   		OWF_Result[4].31:=0;
   		OWF_Result[5]:=OWF_Result[5] + 263129127+OWF_Add_c;
   		OWF_Add_c.5:=OWF_Result[5].31;
   		OWF_Result[5].31:=0;
   		OWF_Result[6]:=OWF_Result[6] + 1259933343+OWF_Add_c;
   		OWF_Add_c.6:=OWF_Result[6].31;
   		OWF_Result[6].31:=0;
   		OWF_Result[7]:=OWF_Result[7] + 1026723117+OWF_Add_c;
   		OWF_Add_c.7:=OWF_Result[7].31;
   		OWF_Result[7].31:=0;
   		OWF_Result[8]:=OWF_Result[8] + 1423999399+OWF_Add_c;
   		OWF_Add_c.8:=OWF_Result[8].31;
   		OWF_Result[8].31:=0;
   	End_If;
   	If OWF_Input[7].[6] Then
   		OWF_Result[0]:=OWF_Result[0] + 1069224909+OWF_Add_c;
   		OWF_Add_c.0:=OWF_Result[0].31;
   		OWF_Result[0].31:=0;
   		OWF_Result[1]:=OWF_Result[1] + 1534942001+OWF_Add_c;
   		OWF_Add_c.1:=OWF_Result[1].31;
   		OWF_Result[1].31:=0;
   		OWF_Result[2]:=OWF_Result[2] + 2056683021+OWF_Add_c;
   		OWF_Add_c.2:=OWF_Result[2].31;
   		OWF_Result[2].31:=0;
   		OWF_Result[3]:=OWF_Result[3] + 1056347500+OWF_Add_c;
   		OWF_Add_c.3:=OWF_Result[3].31;
   		OWF_Result[3].31:=0;
   		OWF_Result[4]:=OWF_Result[4] + 944436856+OWF_Add_c;
   		OWF_Add_c.4:=OWF_Result[4].31;
   		OWF_Result[4].31:=0;
   		OWF_Result[5]:=OWF_Result[5] + 288371840+OWF_Add_c;
   		OWF_Add_c.5:=OWF_Result[5].31;
   		OWF_Result[5].31:=0;
   		OWF_Result[6]:=OWF_Result[6] + 1541197734+OWF_Add_c;
   		OWF_Add_c.6:=OWF_Result[6].31;
   		OWF_Result[6].31:=0;
   		OWF_Result[7]:=OWF_Result[7] + 945574548+OWF_Add_c;
   		OWF_Add_c.7:=OWF_Result[7].31;
   		OWF_Result[7].31:=0;
   		OWF_Result[8]:=OWF_Result[8] + 925934982+OWF_Add_c;
   		OWF_Add_c.8:=OWF_Result[8].31;
   		OWF_Result[8].31:=0;
   	End_If;
   	If OWF_Input[7].[7] Then
   		OWF_Result[0]:=OWF_Result[0] + 2027697593+OWF_Add_c;
   		OWF_Add_c.0:=OWF_Result[0].31;
   		OWF_Result[0].31:=0;
   		OWF_Result[1]:=OWF_Result[1] + 1826137534+OWF_Add_c;
   		OWF_Add_c.1:=OWF_Result[1].31;
   		OWF_Result[1].31:=0;
   		OWF_Result[2]:=OWF_Result[2] + 1291417064+OWF_Add_c;
   		OWF_Add_c.2:=OWF_Result[2].31;
   		OWF_Result[2].31:=0;
   		OWF_Result[3]:=OWF_Result[3] + 1315183552+OWF_Add_c;
   		OWF_Add_c.3:=OWF_Result[3].31;
   		OWF_Result[3].31:=0;
   		OWF_Result[4]:=OWF_Result[4] + 492557432+OWF_Add_c;
   		OWF_Add_c.4:=OWF_Result[4].31;
   		OWF_Result[4].31:=0;
   		OWF_Result[5]:=OWF_Result[5] + 618670102+OWF_Add_c;
   		OWF_Add_c.5:=OWF_Result[5].31;
   		OWF_Result[5].31:=0;
   		OWF_Result[6]:=OWF_Result[6] + 2053349736+OWF_Add_c;
   		OWF_Add_c.6:=OWF_Result[6].31;
   		OWF_Result[6].31:=0;
   		OWF_Result[7]:=OWF_Result[7] + 286016371+OWF_Add_c;
   		OWF_Add_c.7:=OWF_Result[7].31;
   		OWF_Result[7].31:=0;
   		OWF_Result[8]:=OWF_Result[8] + 34477476+OWF_Add_c;
   		OWF_Add_c.8:=OWF_Result[8].31;
   		OWF_Result[8].31:=0;
   	End_If;
   	If OWF_Input[7].[8] Then
   		OWF_Result[0]:=OWF_Result[0] + 1609993904+OWF_Add_c;
   		OWF_Add_c.0:=OWF_Result[0].31;
   		OWF_Result[0].31:=0;
   		OWF_Result[1]:=OWF_Result[1] + 285268351+OWF_Add_c;
   		OWF_Add_c.1:=OWF_Result[1].31;
   		OWF_Result[1].31:=0;
   		OWF_Result[2]:=OWF_Result[2] + 1049093750+OWF_Add_c;
   		OWF_Add_c.2:=OWF_Result[2].31;
   		OWF_Result[2].31:=0;
   		OWF_Result[3]:=OWF_Result[3] + 12994338+OWF_Add_c;
   		OWF_Add_c.3:=OWF_Result[3].31;
   		OWF_Result[3].31:=0;
   		OWF_Result[4]:=OWF_Result[4] + 1664386814+OWF_Add_c;
   		OWF_Add_c.4:=OWF_Result[4].31;
   		OWF_Result[4].31:=0;
   		OWF_Result[5]:=OWF_Result[5] + 1612356757+OWF_Add_c;
   		OWF_Add_c.5:=OWF_Result[5].31;
   		OWF_Result[5].31:=0;
   		OWF_Result[6]:=OWF_Result[6] + 950446094+OWF_Add_c;
   		OWF_Add_c.6:=OWF_Result[6].31;
   		OWF_Result[6].31:=0;
   		OWF_Result[7]:=OWF_Result[7] + 766006761+OWF_Add_c;
   		OWF_Add_c.7:=OWF_Result[7].31;
   		OWF_Result[7].31:=0;
   		OWF_Result[8]:=OWF_Result[8] + 1355626236+OWF_Add_c;
   		OWF_Add_c.8:=OWF_Result[8].31;
   		OWF_Result[8].31:=0;
   	End_If;
   	If OWF_Input[7].[9] Then
   		OWF_Result[0]:=OWF_Result[0] + 694616675+OWF_Add_c;
   		OWF_Add_c.0:=OWF_Result[0].31;
   		OWF_Result[0].31:=0;
   		OWF_Result[1]:=OWF_Result[1] + 1636383722+OWF_Add_c;
   		OWF_Add_c.1:=OWF_Result[1].31;
   		OWF_Result[1].31:=0;
   		OWF_Result[2]:=OWF_Result[2] + 813808724+OWF_Add_c;
   		OWF_Add_c.2:=OWF_Result[2].31;
   		OWF_Result[2].31:=0;
   		OWF_Result[3]:=OWF_Result[3] + 1441798455+OWF_Add_c;
   		OWF_Add_c.3:=OWF_Result[3].31;
   		OWF_Result[3].31:=0;
   		OWF_Result[4]:=OWF_Result[4] + 205766012+OWF_Add_c;
   		OWF_Add_c.4:=OWF_Result[4].31;
   		OWF_Result[4].31:=0;
   		OWF_Result[5]:=OWF_Result[5] + 589639203+OWF_Add_c;
   		OWF_Add_c.5:=OWF_Result[5].31;
   		OWF_Result[5].31:=0;
   		OWF_Result[6]:=OWF_Result[6] + 1829006817+OWF_Add_c;
   		OWF_Add_c.6:=OWF_Result[6].31;
   		OWF_Result[6].31:=0;
   		OWF_Result[7]:=OWF_Result[7] + 1285210054+OWF_Add_c;
   		OWF_Add_c.7:=OWF_Result[7].31;
   		OWF_Result[7].31:=0;
   		OWF_Result[8]:=OWF_Result[8] + 152212693+OWF_Add_c;
   		OWF_Add_c.8:=OWF_Result[8].31;
   		OWF_Result[8].31:=0;
   	End_If;
   	If OWF_Input[7].[10] Then
   		OWF_Result[0]:=OWF_Result[0] + 306590462+OWF_Add_c;
   		OWF_Add_c.0:=OWF_Result[0].31;
   		OWF_Result[0].31:=0;
   		OWF_Result[1]:=OWF_Result[1] + 463214707+OWF_Add_c;
   		OWF_Add_c.1:=OWF_Result[1].31;
   		OWF_Result[1].31:=0;
   		OWF_Result[2]:=OWF_Result[2] + 1073243492+OWF_Add_c;
   		OWF_Add_c.2:=OWF_Result[2].31;
   		OWF_Result[2].31:=0;
   		OWF_Result[3]:=OWF_Result[3] + 1498408871+OWF_Add_c;
   		OWF_Add_c.3:=OWF_Result[3].31;
   		OWF_Result[3].31:=0;
   		OWF_Result[4]:=OWF_Result[4] + 1121005884+OWF_Add_c;
   		OWF_Add_c.4:=OWF_Result[4].31;
   		OWF_Result[4].31:=0;
   		OWF_Result[5]:=OWF_Result[5] + 1933284086+OWF_Add_c;
   		OWF_Add_c.5:=OWF_Result[5].31;
   		OWF_Result[5].31:=0;
   		OWF_Result[6]:=OWF_Result[6] + 1141991459+OWF_Add_c;
   		OWF_Add_c.6:=OWF_Result[6].31;
   		OWF_Result[6].31:=0;
   		OWF_Result[7]:=OWF_Result[7] + 1146716215+OWF_Add_c;
   		OWF_Add_c.7:=OWF_Result[7].31;
   		OWF_Result[7].31:=0;
   		OWF_Result[8]:=OWF_Result[8] + 1107820603+OWF_Add_c;
   		OWF_Add_c.8:=OWF_Result[8].31;
   		OWF_Result[8].31:=0;
   	End_If;
   	If OWF_Input[7].[11] Then
   		OWF_Result[0]:=OWF_Result[0] + 512819892+OWF_Add_c;
   		OWF_Add_c.0:=OWF_Result[0].31;
   		OWF_Result[0].31:=0;
   		OWF_Result[1]:=OWF_Result[1] + 23616385+OWF_Add_c;
   		OWF_Add_c.1:=OWF_Result[1].31;
   		OWF_Result[1].31:=0;
   		OWF_Result[2]:=OWF_Result[2] + 917671887+OWF_Add_c;
   		OWF_Add_c.2:=OWF_Result[2].31;
   		OWF_Result[2].31:=0;
   		OWF_Result[3]:=OWF_Result[3] + 355867720+OWF_Add_c;
   		OWF_Add_c.3:=OWF_Result[3].31;
   		OWF_Result[3].31:=0;
   		OWF_Result[4]:=OWF_Result[4] + 1478009650+OWF_Add_c;
   		OWF_Add_c.4:=OWF_Result[4].31;
   		OWF_Result[4].31:=0;
   		OWF_Result[5]:=OWF_Result[5] + 1568264334+OWF_Add_c;
   		OWF_Add_c.5:=OWF_Result[5].31;
   		OWF_Result[5].31:=0;
   		OWF_Result[6]:=OWF_Result[6] + 1184924613+OWF_Add_c;
   		OWF_Add_c.6:=OWF_Result[6].31;
   		OWF_Result[6].31:=0;
   		OWF_Result[7]:=OWF_Result[7] + 1527868064+OWF_Add_c;
   		OWF_Add_c.7:=OWF_Result[7].31;
   		OWF_Result[7].31:=0;
   		OWF_Result[8]:=OWF_Result[8] + 2072058158+OWF_Add_c;
   		OWF_Add_c.8:=OWF_Result[8].31;
   		OWF_Result[8].31:=0;
   	End_If;
   	If OWF_Input[7].[12] Then
   		OWF_Result[0]:=OWF_Result[0] + 1014625951+OWF_Add_c;
   		OWF_Add_c.0:=OWF_Result[0].31;
   		OWF_Result[0].31:=0;
   		OWF_Result[1]:=OWF_Result[1] + 1533249236+OWF_Add_c;
   		OWF_Add_c.1:=OWF_Result[1].31;
   		OWF_Result[1].31:=0;
   		OWF_Result[2]:=OWF_Result[2] + 2130006381+OWF_Add_c;
   		OWF_Add_c.2:=OWF_Result[2].31;
   		OWF_Result[2].31:=0;
   		OWF_Result[3]:=OWF_Result[3] + 2146846276+OWF_Add_c;
   		OWF_Add_c.3:=OWF_Result[3].31;
   		OWF_Result[3].31:=0;
   		OWF_Result[4]:=OWF_Result[4] + 1646388285+OWF_Add_c;
   		OWF_Add_c.4:=OWF_Result[4].31;
   		OWF_Result[4].31:=0;
   		OWF_Result[5]:=OWF_Result[5] + 1699246205+OWF_Add_c;
   		OWF_Add_c.5:=OWF_Result[5].31;
   		OWF_Result[5].31:=0;
   		OWF_Result[6]:=OWF_Result[6] + 559380684+OWF_Add_c;
   		OWF_Add_c.6:=OWF_Result[6].31;
   		OWF_Result[6].31:=0;
   		OWF_Result[7]:=OWF_Result[7] + 1307307102+OWF_Add_c;
   		OWF_Add_c.7:=OWF_Result[7].31;
   		OWF_Result[7].31:=0;
   		OWF_Result[8]:=OWF_Result[8] + 606704531+OWF_Add_c;
   		OWF_Add_c.8:=OWF_Result[8].31;
   		OWF_Result[8].31:=0;
   	End_If;
   	If OWF_Input[7].[13] Then
   		OWF_Result[0]:=OWF_Result[0] + 1359161121+OWF_Add_c;
   		OWF_Add_c.0:=OWF_Result[0].31;
   		OWF_Result[0].31:=0;
   		OWF_Result[1]:=OWF_Result[1] + 1918952380+OWF_Add_c;
   		OWF_Add_c.1:=OWF_Result[1].31;
   		OWF_Result[1].31:=0;
   		OWF_Result[2]:=OWF_Result[2] + 1473068338+OWF_Add_c;
   		OWF_Add_c.2:=OWF_Result[2].31;
   		OWF_Result[2].31:=0;
   		OWF_Result[3]:=OWF_Result[3] + 1693090892+OWF_Add_c;
   		OWF_Add_c.3:=OWF_Result[3].31;
   		OWF_Result[3].31:=0;
   		OWF_Result[4]:=OWF_Result[4] + 1915525502+OWF_Add_c;
   		OWF_Add_c.4:=OWF_Result[4].31;
   		OWF_Result[4].31:=0;
   		OWF_Result[5]:=OWF_Result[5] + 1372317013+OWF_Add_c;
   		OWF_Add_c.5:=OWF_Result[5].31;
   		OWF_Result[5].31:=0;
   		OWF_Result[6]:=OWF_Result[6] + 99771102+OWF_Add_c;
   		OWF_Add_c.6:=OWF_Result[6].31;
   		OWF_Result[6].31:=0;
   		OWF_Result[7]:=OWF_Result[7] + 192894431+OWF_Add_c;
   		OWF_Add_c.7:=OWF_Result[7].31;
   		OWF_Result[7].31:=0;
   		OWF_Result[8]:=OWF_Result[8] + 1744731961+OWF_Add_c;
   		OWF_Add_c.8:=OWF_Result[8].31;
   		OWF_Result[8].31:=0;
   	End_If;
   	If OWF_Input[7].[14] Then
   		OWF_Result[0]:=OWF_Result[0] + 1706736508+OWF_Add_c;
   		OWF_Add_c.0:=OWF_Result[0].31;
   		OWF_Result[0].31:=0;
   		OWF_Result[1]:=OWF_Result[1] + 1484877150+OWF_Add_c;
   		OWF_Add_c.1:=OWF_Result[1].31;
   		OWF_Result[1].31:=0;
   		OWF_Result[2]:=OWF_Result[2] + 869604235+OWF_Add_c;
   		OWF_Add_c.2:=OWF_Result[2].31;
   		OWF_Result[2].31:=0;
   		OWF_Result[3]:=OWF_Result[3] + 1353356392+OWF_Add_c;
   		OWF_Add_c.3:=OWF_Result[3].31;
   		OWF_Result[3].31:=0;
   		OWF_Result[4]:=OWF_Result[4] + 347447568+OWF_Add_c;
   		OWF_Add_c.4:=OWF_Result[4].31;
   		OWF_Result[4].31:=0;
   		OWF_Result[5]:=OWF_Result[5] + 1293208581+OWF_Add_c;
   		OWF_Add_c.5:=OWF_Result[5].31;
   		OWF_Result[5].31:=0;
   		OWF_Result[6]:=OWF_Result[6] + 1575776397+OWF_Add_c;
   		OWF_Add_c.6:=OWF_Result[6].31;
   		OWF_Result[6].31:=0;
   		OWF_Result[7]:=OWF_Result[7] + 1427687325+OWF_Add_c;
   		OWF_Add_c.7:=OWF_Result[7].31;
   		OWF_Result[7].31:=0;
   		OWF_Result[8]:=OWF_Result[8] + 935165463+OWF_Add_c;
   		OWF_Add_c.8:=OWF_Result[8].31;
   		OWF_Result[8].31:=0;
   	End_If;
   	If OWF_Input[7].[15] Then
   		OWF_Result[0]:=OWF_Result[0] + 1743664197+OWF_Add_c;
   		OWF_Add_c.0:=OWF_Result[0].31;
   		OWF_Result[0].31:=0;
   		OWF_Result[1]:=OWF_Result[1] + 706528617+OWF_Add_c;
   		OWF_Add_c.1:=OWF_Result[1].31;
   		OWF_Result[1].31:=0;
   		OWF_Result[2]:=OWF_Result[2] + 1958351723+OWF_Add_c;
   		OWF_Add_c.2:=OWF_Result[2].31;
   		OWF_Result[2].31:=0;
   		OWF_Result[3]:=OWF_Result[3] + 82257141+OWF_Add_c;
   		OWF_Add_c.3:=OWF_Result[3].31;
   		OWF_Result[3].31:=0;
   		OWF_Result[4]:=OWF_Result[4] + 860284908+OWF_Add_c;
   		OWF_Add_c.4:=OWF_Result[4].31;
   		OWF_Result[4].31:=0;
   		OWF_Result[5]:=OWF_Result[5] + 1587356663+OWF_Add_c;
   		OWF_Add_c.5:=OWF_Result[5].31;
   		OWF_Result[5].31:=0;
   		OWF_Result[6]:=OWF_Result[6] + 1299103155+OWF_Add_c;
   		OWF_Add_c.6:=OWF_Result[6].31;
   		OWF_Result[6].31:=0;
   		OWF_Result[7]:=OWF_Result[7] + 1945550030+OWF_Add_c;
   		OWF_Add_c.7:=OWF_Result[7].31;
   		OWF_Result[7].31:=0;
   		OWF_Result[8]:=OWF_Result[8] + 2117411835+OWF_Add_c;
   		OWF_Add_c.8:=OWF_Result[8].31;
   		OWF_Result[8].31:=0;
   	End_If;
   	If OWF_Input[7].[16] Then
   		OWF_Result[0]:=OWF_Result[0] + 1713469729+OWF_Add_c;
   		OWF_Add_c.0:=OWF_Result[0].31;
   		OWF_Result[0].31:=0;
   		OWF_Result[1]:=OWF_Result[1] + 581994065+OWF_Add_c;
   		OWF_Add_c.1:=OWF_Result[1].31;
   		OWF_Result[1].31:=0;
   		OWF_Result[2]:=OWF_Result[2] + 190604491+OWF_Add_c;
   		OWF_Add_c.2:=OWF_Result[2].31;
   		OWF_Result[2].31:=0;
   		OWF_Result[3]:=OWF_Result[3] + 1975804182+OWF_Add_c;
   		OWF_Add_c.3:=OWF_Result[3].31;
   		OWF_Result[3].31:=0;
   		OWF_Result[4]:=OWF_Result[4] + 1579426154+OWF_Add_c;
   		OWF_Add_c.4:=OWF_Result[4].31;
   		OWF_Result[4].31:=0;
   		OWF_Result[5]:=OWF_Result[5] + 1526883195+OWF_Add_c;
   		OWF_Add_c.5:=OWF_Result[5].31;
   		OWF_Result[5].31:=0;
   		OWF_Result[6]:=OWF_Result[6] + 1534112395+OWF_Add_c;
   		OWF_Add_c.6:=OWF_Result[6].31;
   		OWF_Result[6].31:=0;
   		OWF_Result[7]:=OWF_Result[7] + 1953195996+OWF_Add_c;
   		OWF_Add_c.7:=OWF_Result[7].31;
   		OWF_Result[7].31:=0;
   		OWF_Result[8]:=OWF_Result[8] + 1196776541+OWF_Add_c;
   		OWF_Add_c.8:=OWF_Result[8].31;
   		OWF_Result[8].31:=0;
   	End_If;
   	If OWF_Input[7].[17] Then
   		OWF_Result[0]:=OWF_Result[0] + 1352341478+OWF_Add_c;
   		OWF_Add_c.0:=OWF_Result[0].31;
   		OWF_Result[0].31:=0;
   		OWF_Result[1]:=OWF_Result[1] + 1327190218+OWF_Add_c;
   		OWF_Add_c.1:=OWF_Result[1].31;
   		OWF_Result[1].31:=0;
   		OWF_Result[2]:=OWF_Result[2] + 1940036231+OWF_Add_c;
   		OWF_Add_c.2:=OWF_Result[2].31;
   		OWF_Result[2].31:=0;
   		OWF_Result[3]:=OWF_Result[3] + 569828080+OWF_Add_c;
   		OWF_Add_c.3:=OWF_Result[3].31;
   		OWF_Result[3].31:=0;
   		OWF_Result[4]:=OWF_Result[4] + 1243727683+OWF_Add_c;
   		OWF_Add_c.4:=OWF_Result[4].31;
   		OWF_Result[4].31:=0;
   		OWF_Result[5]:=OWF_Result[5] + 741960146+OWF_Add_c;
   		OWF_Add_c.5:=OWF_Result[5].31;
   		OWF_Result[5].31:=0;
   		OWF_Result[6]:=OWF_Result[6] + 2046665451+OWF_Add_c;
   		OWF_Add_c.6:=OWF_Result[6].31;
   		OWF_Result[6].31:=0;
   		OWF_Result[7]:=OWF_Result[7] + 482388128+OWF_Add_c;
   		OWF_Add_c.7:=OWF_Result[7].31;
   		OWF_Result[7].31:=0;
   		OWF_Result[8]:=OWF_Result[8] + 1415487699+OWF_Add_c;
   		OWF_Add_c.8:=OWF_Result[8].31;
   		OWF_Result[8].31:=0;
   	End_If;
   	If OWF_Input[7].[18] Then
   		OWF_Result[0]:=OWF_Result[0] + 419967488+OWF_Add_c;
   		OWF_Add_c.0:=OWF_Result[0].31;
   		OWF_Result[0].31:=0;
   		OWF_Result[1]:=OWF_Result[1] + 319301420+OWF_Add_c;
   		OWF_Add_c.1:=OWF_Result[1].31;
   		OWF_Result[1].31:=0;
   		OWF_Result[2]:=OWF_Result[2] + 1439251767+OWF_Add_c;
   		OWF_Add_c.2:=OWF_Result[2].31;
   		OWF_Result[2].31:=0;
   		OWF_Result[3]:=OWF_Result[3] + 159030407+OWF_Add_c;
   		OWF_Add_c.3:=OWF_Result[3].31;
   		OWF_Result[3].31:=0;
   		OWF_Result[4]:=OWF_Result[4] + 1688057992+OWF_Add_c;
   		OWF_Add_c.4:=OWF_Result[4].31;
   		OWF_Result[4].31:=0;
   		OWF_Result[5]:=OWF_Result[5] + 677856544+OWF_Add_c;
   		OWF_Add_c.5:=OWF_Result[5].31;
   		OWF_Result[5].31:=0;
   		OWF_Result[6]:=OWF_Result[6] + 1921290271+OWF_Add_c;
   		OWF_Add_c.6:=OWF_Result[6].31;
   		OWF_Result[6].31:=0;
   		OWF_Result[7]:=OWF_Result[7] + 1347176510+OWF_Add_c;
   		OWF_Add_c.7:=OWF_Result[7].31;
   		OWF_Result[7].31:=0;
   		OWF_Result[8]:=OWF_Result[8] + 1129087746+OWF_Add_c;
   		OWF_Add_c.8:=OWF_Result[8].31;
   		OWF_Result[8].31:=0;
   	End_If;
   	If OWF_Input[7].[19] Then
   		OWF_Result[0]:=OWF_Result[0] + 909989480+OWF_Add_c;
   		OWF_Add_c.0:=OWF_Result[0].31;
   		OWF_Result[0].31:=0;
   		OWF_Result[1]:=OWF_Result[1] + 70607674+OWF_Add_c;
   		OWF_Add_c.1:=OWF_Result[1].31;
   		OWF_Result[1].31:=0;
   		OWF_Result[2]:=OWF_Result[2] + 102357735+OWF_Add_c;
   		OWF_Add_c.2:=OWF_Result[2].31;
   		OWF_Result[2].31:=0;
   		OWF_Result[3]:=OWF_Result[3] + 1548947751+OWF_Add_c;
   		OWF_Add_c.3:=OWF_Result[3].31;
   		OWF_Result[3].31:=0;
   		OWF_Result[4]:=OWF_Result[4] + 1541273950+OWF_Add_c;
   		OWF_Add_c.4:=OWF_Result[4].31;
   		OWF_Result[4].31:=0;
   		OWF_Result[5]:=OWF_Result[5] + 1965581916+OWF_Add_c;
   		OWF_Add_c.5:=OWF_Result[5].31;
   		OWF_Result[5].31:=0;
   		OWF_Result[6]:=OWF_Result[6] + 714783171+OWF_Add_c;
   		OWF_Add_c.6:=OWF_Result[6].31;
   		OWF_Result[6].31:=0;
   		OWF_Result[7]:=OWF_Result[7] + 952638591+OWF_Add_c;
   		OWF_Add_c.7:=OWF_Result[7].31;
   		OWF_Result[7].31:=0;
   		OWF_Result[8]:=OWF_Result[8] + 1892750752+OWF_Add_c;
   		OWF_Add_c.8:=OWF_Result[8].31;
   		OWF_Result[8].31:=0;
   	End_If;
   	If OWF_Input[7].[20] Then
   		OWF_Result[0]:=OWF_Result[0] + 1923601846+OWF_Add_c;
   		OWF_Add_c.0:=OWF_Result[0].31;
   		OWF_Result[0].31:=0;
   		OWF_Result[1]:=OWF_Result[1] + 431367542+OWF_Add_c;
   		OWF_Add_c.1:=OWF_Result[1].31;
   		OWF_Result[1].31:=0;
   		OWF_Result[2]:=OWF_Result[2] + 812772690+OWF_Add_c;
   		OWF_Add_c.2:=OWF_Result[2].31;
   		OWF_Result[2].31:=0;
   		OWF_Result[3]:=OWF_Result[3] + 1612004830+OWF_Add_c;
   		OWF_Add_c.3:=OWF_Result[3].31;
   		OWF_Result[3].31:=0;
   		OWF_Result[4]:=OWF_Result[4] + 1503607425+OWF_Add_c;
   		OWF_Add_c.4:=OWF_Result[4].31;
   		OWF_Result[4].31:=0;
   		OWF_Result[5]:=OWF_Result[5] + 257117095+OWF_Add_c;
   		OWF_Add_c.5:=OWF_Result[5].31;
   		OWF_Result[5].31:=0;
   		OWF_Result[6]:=OWF_Result[6] + 1165565758+OWF_Add_c;
   		OWF_Add_c.6:=OWF_Result[6].31;
   		OWF_Result[6].31:=0;
   		OWF_Result[7]:=OWF_Result[7] + 1791078952+OWF_Add_c;
   		OWF_Add_c.7:=OWF_Result[7].31;
   		OWF_Result[7].31:=0;
   		OWF_Result[8]:=OWF_Result[8] + 1316586480+OWF_Add_c;
   		OWF_Add_c.8:=OWF_Result[8].31;
   		OWF_Result[8].31:=0;
   	End_If;
   	If OWF_Input[7].[21] Then
   		OWF_Result[0]:=OWF_Result[0] + 1179130031+OWF_Add_c;
   		OWF_Add_c.0:=OWF_Result[0].31;
   		OWF_Result[0].31:=0;
   		OWF_Result[1]:=OWF_Result[1] + 1413483742+OWF_Add_c;
   		OWF_Add_c.1:=OWF_Result[1].31;
   		OWF_Result[1].31:=0;
   		OWF_Result[2]:=OWF_Result[2] + 2076538493+OWF_Add_c;
   		OWF_Add_c.2:=OWF_Result[2].31;
   		OWF_Result[2].31:=0;
   		OWF_Result[3]:=OWF_Result[3] + 415974763+OWF_Add_c;
   		OWF_Add_c.3:=OWF_Result[3].31;
   		OWF_Result[3].31:=0;
   		OWF_Result[4]:=OWF_Result[4] + 461079233+OWF_Add_c;
   		OWF_Add_c.4:=OWF_Result[4].31;
   		OWF_Result[4].31:=0;
   		OWF_Result[5]:=OWF_Result[5] + 207770264+OWF_Add_c;
   		OWF_Add_c.5:=OWF_Result[5].31;
   		OWF_Result[5].31:=0;
   		OWF_Result[6]:=OWF_Result[6] + 670532004+OWF_Add_c;
   		OWF_Add_c.6:=OWF_Result[6].31;
   		OWF_Result[6].31:=0;
   		OWF_Result[7]:=OWF_Result[7] + 164283060+OWF_Add_c;
   		OWF_Add_c.7:=OWF_Result[7].31;
   		OWF_Result[7].31:=0;
   		OWF_Result[8]:=OWF_Result[8] + 1512816438+OWF_Add_c;
   		OWF_Add_c.8:=OWF_Result[8].31;
   		OWF_Result[8].31:=0;
   	End_If;
   	If OWF_Input[7].[22] Then
   		OWF_Result[0]:=OWF_Result[0] + 1897360171+OWF_Add_c;
   		OWF_Add_c.0:=OWF_Result[0].31;
   		OWF_Result[0].31:=0;
   		OWF_Result[1]:=OWF_Result[1] + 1308779824+OWF_Add_c;
   		OWF_Add_c.1:=OWF_Result[1].31;
   		OWF_Result[1].31:=0;
   		OWF_Result[2]:=OWF_Result[2] + 1875593423+OWF_Add_c;
   		OWF_Add_c.2:=OWF_Result[2].31;
   		OWF_Result[2].31:=0;
   		OWF_Result[3]:=OWF_Result[3] + 571271217+OWF_Add_c;
   		OWF_Add_c.3:=OWF_Result[3].31;
   		OWF_Result[3].31:=0;
   		OWF_Result[4]:=OWF_Result[4] + 344940971+OWF_Add_c;
   		OWF_Add_c.4:=OWF_Result[4].31;
   		OWF_Result[4].31:=0;
   		OWF_Result[5]:=OWF_Result[5] + 75339231+OWF_Add_c;
   		OWF_Add_c.5:=OWF_Result[5].31;
   		OWF_Result[5].31:=0;
   		OWF_Result[6]:=OWF_Result[6] + 1428316860+OWF_Add_c;
   		OWF_Add_c.6:=OWF_Result[6].31;
   		OWF_Result[6].31:=0;
   		OWF_Result[7]:=OWF_Result[7] + 1811603075+OWF_Add_c;
   		OWF_Add_c.7:=OWF_Result[7].31;
   		OWF_Result[7].31:=0;
   		OWF_Result[8]:=OWF_Result[8] + 1679786029+OWF_Add_c;
   		OWF_Add_c.8:=OWF_Result[8].31;
   		OWF_Result[8].31:=0;
   	End_If;
   	If OWF_Input[7].[23] Then
   		OWF_Result[0]:=OWF_Result[0] + 271831917+OWF_Add_c;
   		OWF_Add_c.0:=OWF_Result[0].31;
   		OWF_Result[0].31:=0;
   		OWF_Result[1]:=OWF_Result[1] + 663117307+OWF_Add_c;
   		OWF_Add_c.1:=OWF_Result[1].31;
   		OWF_Result[1].31:=0;
   		OWF_Result[2]:=OWF_Result[2] + 1802435718+OWF_Add_c;
   		OWF_Add_c.2:=OWF_Result[2].31;
   		OWF_Result[2].31:=0;
   		OWF_Result[3]:=OWF_Result[3] + 585874673+OWF_Add_c;
   		OWF_Add_c.3:=OWF_Result[3].31;
   		OWF_Result[3].31:=0;
   		OWF_Result[4]:=OWF_Result[4] + 701698092+OWF_Add_c;
   		OWF_Add_c.4:=OWF_Result[4].31;
   		OWF_Result[4].31:=0;
   		OWF_Result[5]:=OWF_Result[5] + 1402770880+OWF_Add_c;
   		OWF_Add_c.5:=OWF_Result[5].31;
   		OWF_Result[5].31:=0;
   		OWF_Result[6]:=OWF_Result[6] + 452824658+OWF_Add_c;
   		OWF_Add_c.6:=OWF_Result[6].31;
   		OWF_Result[6].31:=0;
   		OWF_Result[7]:=OWF_Result[7] + 1400742763+OWF_Add_c;
   		OWF_Add_c.7:=OWF_Result[7].31;
   		OWF_Result[7].31:=0;
   		OWF_Result[8]:=OWF_Result[8] + 2073024045+OWF_Add_c;
   		OWF_Add_c.8:=OWF_Result[8].31;
   		OWF_Result[8].31:=0;
   	End_If;
   	If OWF_Input[7].[24] Then
   		OWF_Result[0]:=OWF_Result[0] + 1367845667+OWF_Add_c;
   		OWF_Add_c.0:=OWF_Result[0].31;
   		OWF_Result[0].31:=0;
   		OWF_Result[1]:=OWF_Result[1] + 1195094582+OWF_Add_c;
   		OWF_Add_c.1:=OWF_Result[1].31;
   		OWF_Result[1].31:=0;
   		OWF_Result[2]:=OWF_Result[2] + 494736933+OWF_Add_c;
   		OWF_Add_c.2:=OWF_Result[2].31;
   		OWF_Result[2].31:=0;
   		OWF_Result[3]:=OWF_Result[3] + 1875737261+OWF_Add_c;
   		OWF_Add_c.3:=OWF_Result[3].31;
   		OWF_Result[3].31:=0;
   		OWF_Result[4]:=OWF_Result[4] + 726339725+OWF_Add_c;
   		OWF_Add_c.4:=OWF_Result[4].31;
   		OWF_Result[4].31:=0;
   		OWF_Result[5]:=OWF_Result[5] + 1862851936+OWF_Add_c;
   		OWF_Add_c.5:=OWF_Result[5].31;
   		OWF_Result[5].31:=0;
   		OWF_Result[6]:=OWF_Result[6] + 296798862+OWF_Add_c;
   		OWF_Add_c.6:=OWF_Result[6].31;
   		OWF_Result[6].31:=0;
   		OWF_Result[7]:=OWF_Result[7] + 1485306441+OWF_Add_c;
   		OWF_Add_c.7:=OWF_Result[7].31;
   		OWF_Result[7].31:=0;
   		OWF_Result[8]:=OWF_Result[8] + 79244469+OWF_Add_c;
   		OWF_Add_c.8:=OWF_Result[8].31;
   		OWF_Result[8].31:=0;
   	End_If;
   	If OWF_Input[7].[25] Then
   		OWF_Result[0]:=OWF_Result[0] + 1748009068+OWF_Add_c;
   		OWF_Add_c.0:=OWF_Result[0].31;
   		OWF_Result[0].31:=0;
   		OWF_Result[1]:=OWF_Result[1] + 153673379+OWF_Add_c;
   		OWF_Add_c.1:=OWF_Result[1].31;
   		OWF_Result[1].31:=0;
   		OWF_Result[2]:=OWF_Result[2] + 1563899973+OWF_Add_c;
   		OWF_Add_c.2:=OWF_Result[2].31;
   		OWF_Result[2].31:=0;
   		OWF_Result[3]:=OWF_Result[3] + 210477071+OWF_Add_c;
   		OWF_Add_c.3:=OWF_Result[3].31;
   		OWF_Result[3].31:=0;
   		OWF_Result[4]:=OWF_Result[4] + 598591903+OWF_Add_c;
   		OWF_Add_c.4:=OWF_Result[4].31;
   		OWF_Result[4].31:=0;
   		OWF_Result[5]:=OWF_Result[5] + 889903791+OWF_Add_c;
   		OWF_Add_c.5:=OWF_Result[5].31;
   		OWF_Result[5].31:=0;
   		OWF_Result[6]:=OWF_Result[6] + 1087681228+OWF_Add_c;
   		OWF_Add_c.6:=OWF_Result[6].31;
   		OWF_Result[6].31:=0;
   		OWF_Result[7]:=OWF_Result[7] + 146945819+OWF_Add_c;
   		OWF_Add_c.7:=OWF_Result[7].31;
   		OWF_Result[7].31:=0;
   		OWF_Result[8]:=OWF_Result[8] + 658778953+OWF_Add_c;
   		OWF_Add_c.8:=OWF_Result[8].31;
   		OWF_Result[8].31:=0;
   	End_If;
   	If OWF_Input[7].[26] Then
   		OWF_Result[0]:=OWF_Result[0] + 1388889236+OWF_Add_c;
   		OWF_Add_c.0:=OWF_Result[0].31;
   		OWF_Result[0].31:=0;
   		OWF_Result[1]:=OWF_Result[1] + 1854230592+OWF_Add_c;
   		OWF_Add_c.1:=OWF_Result[1].31;
   		OWF_Result[1].31:=0;
   		OWF_Result[2]:=OWF_Result[2] + 1952659775+OWF_Add_c;
   		OWF_Add_c.2:=OWF_Result[2].31;
   		OWF_Result[2].31:=0;
   		OWF_Result[3]:=OWF_Result[3] + 693016622+OWF_Add_c;
   		OWF_Add_c.3:=OWF_Result[3].31;
   		OWF_Result[3].31:=0;
   		OWF_Result[4]:=OWF_Result[4] + 19961190+OWF_Add_c;
   		OWF_Add_c.4:=OWF_Result[4].31;
   		OWF_Result[4].31:=0;
   		OWF_Result[5]:=OWF_Result[5] + 1155238848+OWF_Add_c;
   		OWF_Add_c.5:=OWF_Result[5].31;
   		OWF_Result[5].31:=0;
   		OWF_Result[6]:=OWF_Result[6] + 1721973623+OWF_Add_c;
   		OWF_Add_c.6:=OWF_Result[6].31;
   		OWF_Result[6].31:=0;
   		OWF_Result[7]:=OWF_Result[7] + 1298626904+OWF_Add_c;
   		OWF_Add_c.7:=OWF_Result[7].31;
   		OWF_Result[7].31:=0;
   		OWF_Result[8]:=OWF_Result[8] + 704184103+OWF_Add_c;
   		OWF_Add_c.8:=OWF_Result[8].31;
   		OWF_Result[8].31:=0;
   	End_If;
   	If OWF_Input[7].[27] Then
   		OWF_Result[0]:=OWF_Result[0] + 1064559134+OWF_Add_c;
   		OWF_Add_c.0:=OWF_Result[0].31;
   		OWF_Result[0].31:=0;
   		OWF_Result[1]:=OWF_Result[1] + 628496468+OWF_Add_c;
   		OWF_Add_c.1:=OWF_Result[1].31;
   		OWF_Result[1].31:=0;
   		OWF_Result[2]:=OWF_Result[2] + 1741787667+OWF_Add_c;
   		OWF_Add_c.2:=OWF_Result[2].31;
   		OWF_Result[2].31:=0;
   		OWF_Result[3]:=OWF_Result[3] + 650880797+OWF_Add_c;
   		OWF_Add_c.3:=OWF_Result[3].31;
   		OWF_Result[3].31:=0;
   		OWF_Result[4]:=OWF_Result[4] + 927193641+OWF_Add_c;
   		OWF_Add_c.4:=OWF_Result[4].31;
   		OWF_Result[4].31:=0;
   		OWF_Result[5]:=OWF_Result[5] + 690779087+OWF_Add_c;
   		OWF_Add_c.5:=OWF_Result[5].31;
   		OWF_Result[5].31:=0;
   		OWF_Result[6]:=OWF_Result[6] + 1387171811+OWF_Add_c;
   		OWF_Add_c.6:=OWF_Result[6].31;
   		OWF_Result[6].31:=0;
   		OWF_Result[7]:=OWF_Result[7] + 1642242275+OWF_Add_c;
   		OWF_Add_c.7:=OWF_Result[7].31;
   		OWF_Result[7].31:=0;
   		OWF_Result[8]:=OWF_Result[8] + 750154437+OWF_Add_c;
   		OWF_Add_c.8:=OWF_Result[8].31;
   		OWF_Result[8].31:=0;
   	End_If;
   	If OWF_Input[7].[28] Then
   		OWF_Result[0]:=OWF_Result[0] + 1648370074+OWF_Add_c;
   		OWF_Add_c.0:=OWF_Result[0].31;
   		OWF_Result[0].31:=0;
   		OWF_Result[1]:=OWF_Result[1] + 242619355+OWF_Add_c;
   		OWF_Add_c.1:=OWF_Result[1].31;
   		OWF_Result[1].31:=0;
   		OWF_Result[2]:=OWF_Result[2] + 1874736599+OWF_Add_c;
   		OWF_Add_c.2:=OWF_Result[2].31;
   		OWF_Result[2].31:=0;
   		OWF_Result[3]:=OWF_Result[3] + 1413909693+OWF_Add_c;
   		OWF_Add_c.3:=OWF_Result[3].31;
   		OWF_Result[3].31:=0;
   		OWF_Result[4]:=OWF_Result[4] + 415302371+OWF_Add_c;
   		OWF_Add_c.4:=OWF_Result[4].31;
   		OWF_Result[4].31:=0;
   		OWF_Result[5]:=OWF_Result[5] + 2103173316+OWF_Add_c;
   		OWF_Add_c.5:=OWF_Result[5].31;
   		OWF_Result[5].31:=0;
   		OWF_Result[6]:=OWF_Result[6] + 317087375+OWF_Add_c;
   		OWF_Add_c.6:=OWF_Result[6].31;
   		OWF_Result[6].31:=0;
   		OWF_Result[7]:=OWF_Result[7] + 1550821217+OWF_Add_c;
   		OWF_Add_c.7:=OWF_Result[7].31;
   		OWF_Result[7].31:=0;
   		OWF_Result[8]:=OWF_Result[8] + 61155956+OWF_Add_c;
   		OWF_Add_c.8:=OWF_Result[8].31;
   		OWF_Result[8].31:=0;
   	End_If;
   	If OWF_Input[7].[29] Then
   		OWF_Result[0]:=OWF_Result[0] + 632604897+OWF_Add_c;
   		OWF_Add_c.0:=OWF_Result[0].31;
   		OWF_Result[0].31:=0;
   		OWF_Result[1]:=OWF_Result[1] + 1890179507+OWF_Add_c;
   		OWF_Add_c.1:=OWF_Result[1].31;
   		OWF_Result[1].31:=0;
   		OWF_Result[2]:=OWF_Result[2] + 1607995656+OWF_Add_c;
   		OWF_Add_c.2:=OWF_Result[2].31;
   		OWF_Result[2].31:=0;
   		OWF_Result[3]:=OWF_Result[3] + 1449206150+OWF_Add_c;
   		OWF_Add_c.3:=OWF_Result[3].31;
   		OWF_Result[3].31:=0;
   		OWF_Result[4]:=OWF_Result[4] + 402726737+OWF_Add_c;
   		OWF_Add_c.4:=OWF_Result[4].31;
   		OWF_Result[4].31:=0;
   		OWF_Result[5]:=OWF_Result[5] + 365091023+OWF_Add_c;
   		OWF_Add_c.5:=OWF_Result[5].31;
   		OWF_Result[5].31:=0;
   		OWF_Result[6]:=OWF_Result[6] + 1662601056+OWF_Add_c;
   		OWF_Add_c.6:=OWF_Result[6].31;
   		OWF_Result[6].31:=0;
   		OWF_Result[7]:=OWF_Result[7] + 1022070658+OWF_Add_c;
   		OWF_Add_c.7:=OWF_Result[7].31;
   		OWF_Result[7].31:=0;
   		OWF_Result[8]:=OWF_Result[8] + 49749052+OWF_Add_c;
   		OWF_Add_c.8:=OWF_Result[8].31;
   		OWF_Result[8].31:=0;
   	End_If;
   	If OWF_Input[7].[30] Then
   		OWF_Result[0]:=OWF_Result[0] + 1218340763+OWF_Add_c;
   		OWF_Add_c.0:=OWF_Result[0].31;
   		OWF_Result[0].31:=0;
   		OWF_Result[1]:=OWF_Result[1] + 1701757107+OWF_Add_c;
   		OWF_Add_c.1:=OWF_Result[1].31;
   		OWF_Result[1].31:=0;
   		OWF_Result[2]:=OWF_Result[2] + 1789117076+OWF_Add_c;
   		OWF_Add_c.2:=OWF_Result[2].31;
   		OWF_Result[2].31:=0;
   		OWF_Result[3]:=OWF_Result[3] + 963840108+OWF_Add_c;
   		OWF_Add_c.3:=OWF_Result[3].31;
   		OWF_Result[3].31:=0;
   		OWF_Result[4]:=OWF_Result[4] + 660620140+OWF_Add_c;
   		OWF_Add_c.4:=OWF_Result[4].31;
   		OWF_Result[4].31:=0;
   		OWF_Result[5]:=OWF_Result[5] + 983419398+OWF_Add_c;
   		OWF_Add_c.5:=OWF_Result[5].31;
   		OWF_Result[5].31:=0;
   		OWF_Result[6]:=OWF_Result[6] + 540791099+OWF_Add_c;
   		OWF_Add_c.6:=OWF_Result[6].31;
   		OWF_Result[6].31:=0;
   		OWF_Result[7]:=OWF_Result[7] + 2120149871+OWF_Add_c;
   		OWF_Add_c.7:=OWF_Result[7].31;
   		OWF_Result[7].31:=0;
   		OWF_Result[8]:=OWF_Result[8] + 1356988421+OWF_Add_c;
   		OWF_Add_c.8:=OWF_Result[8].31;
   		OWF_Result[8].31:=0;
   	End_If;
   	If OWF_Input[7].[31] Then
   		OWF_Result[0]:=OWF_Result[0] + 1135594880+OWF_Add_c;
   		OWF_Add_c.0:=OWF_Result[0].31;
   		OWF_Result[0].31:=0;
   		OWF_Result[1]:=OWF_Result[1] + 1430344149+OWF_Add_c;
   		OWF_Add_c.1:=OWF_Result[1].31;
   		OWF_Result[1].31:=0;
   		OWF_Result[2]:=OWF_Result[2] + 426577698+OWF_Add_c;
   		OWF_Add_c.2:=OWF_Result[2].31;
   		OWF_Result[2].31:=0;
   		OWF_Result[3]:=OWF_Result[3] + 34487438+OWF_Add_c;
   		OWF_Add_c.3:=OWF_Result[3].31;
   		OWF_Result[3].31:=0;
   		OWF_Result[4]:=OWF_Result[4] + 142555847+OWF_Add_c;
   		OWF_Add_c.4:=OWF_Result[4].31;
   		OWF_Result[4].31:=0;
   		OWF_Result[5]:=OWF_Result[5] + 380868128+OWF_Add_c;
   		OWF_Add_c.5:=OWF_Result[5].31;
   		OWF_Result[5].31:=0;
   		OWF_Result[6]:=OWF_Result[6] + 797337152+OWF_Add_c;
   		OWF_Add_c.6:=OWF_Result[6].31;
   		OWF_Result[6].31:=0;
   		OWF_Result[7]:=OWF_Result[7] + 1153550956+OWF_Add_c;
   		OWF_Add_c.7:=OWF_Result[7].31;
   		OWF_Result[7].31:=0;
   		OWF_Result[8]:=OWF_Result[8] + 2080693926+OWF_Add_c;
   		OWF_Add_c.8:=OWF_Result[8].31;
   		OWF_Result[8].31:=0;
   	End_If;
   
   	OWF_Result[OWF_InputMaxInd]:=OWF_Result[OWF_InputMaxInd] and 16#FF; //clear high bit
   
END_ROUTINE
